// TIA Portal project "Energy_Drink_V15.1" (V15.1) (continued)
REGION Network 3: *****************************MIXER VALVE********************************************/
         A     "Var_System_DB".Sirupe_Valve.Vlv_Open_Cmd;
         =     "Sirupe_Vlv_Man";

         A     "Var_System_DB".Water_Valve.Vlv_Open_Cmd;
         =     "Water_Vlv_Man";

         A     "Var_System_DB".Tk104_MIXER.Open_Vlv_Cmd;
         O     "HMI_VAR".Man_Valves.Mixer_Discharge_Vlv;
         =     "Mixer_Dis_Vlv";

         A     "Var_System_DB".Cleanning_Process.Vlv_Open_Cmd;
         =     "Mixer_Cleanning_Vlv";
END_REGION

REGION Network 4: *****************************CONVEYOR********************************************/
   // CONVEYOR MAIN CONTACTOR
         A     "Var_System_DB".Conveyor_Belt.M_Main;
         =     "KM1_Main";

   // CONVEYOR STAR CONTACTOR
         A     "Var_System_DB".Conveyor_Belt.M_Star;
         =     "KM2_Star";

   // CONVEYOR DELTA CONTACTOR
         A     "Var_System_DB".Conveyor_Belt.M_Led_Delta;
         =     "KM3_Delta";
END_REGION

REGION Network 5: *******************************PROCESS LEDS****************************************/
   // CONVEYOR BELT MOTOR LED ACTIVATION
         A     "Var_System_DB".Conveyor_Belt.M_Led_Main;
         =     "H4";

         A     "Var_System_DB".Conveyor_Belt.M_Led_Delta;
         =     "H5";

         A     "Var_System_DB".Conveyor_Belt.M_Led_Stop;
         =     "H10";

         A     "Var_System_DB".Conveyor_Belt.M_Led_Ovl;
         =     "H8";

   // MIXER MOTOR LED ACTIVATION
         A     "Var_System_DB".Mixer_Motor.Acel_Led;
         =     "H6";

         A     "Var_System_DB".Mixer_Motor.Decel_Led;
         =     "H7";

         A     "Var_System_DB".Mixer_Motor.Led_Ovl;
         =     "H9";
END_REGION
END_FUNCTION

// folder: 02-START-STOP MANGAMENT

FUNCTION "GENERIC_START-STOP" : Void   // FC1, STL
{ S7_Optimized_Access := 'FALSE' }
VERSION : 0.1
BEGIN

REGION Network 1: ******************************* AUTO MODE ********************************************
   // IF START BUTTON PRESSED => DB START
         A     "Start_Button";
         O     "HMI_VAR".Act_System;
         =     "Var_System_DB".System_Generic.Start;

   // IF DB START ACTIVATED => SYSTEM IS ON
         A     "Var_System_DB".System_Generic.Start;
         AN    "Var_System_DB".System_Generic."Auto/Man";
         FP    "Tag_8";
         S     "Var_System_DB".System_Generic.System_Act;
         S     "Var_System_DB".Conveyor_Belt.M_Stop;

   // IF NEGATIVE EDGE OF DB START => RESET
         A     "Var_System_DB".System_Generic.Start;
         FN    "Tag_9";
         R     "Var_System_DB".System_Generic.Stop_Process;
END_REGION

REGION Network 2: ******************************* MANUAL MODE ********************************************
   // SET MANUAL MODE AUTO/MANUAL = 1
         A     "Var_System_DB".System_Generic."Auto/Man";
         A     "Var_System_DB".System_Generic.Start;
         S     "Var_System_DB".System_Generic.Man_Mode;

   // RESET MANUAL MODE
         AN    "Var_System_DB".System_Generic."Auto/Man";
         R     "Var_System_DB".System_Generic.Man_Mode;
END_REGION

REGION Network 3: ******************************* STOP MODE ********************************************
   // WHILE SYSTEM STOP
         A     "Stop_Button";
         A     "HMI_VAR".Stop_System;
         =     "Var_System_DB".System_Generic.Stop;

         AN    "Stop_Button";
         ON    "HMI_VAR".Stop_System;
         S     "Var_System_DB".System_Generic.Stop_Process;
END_REGION
END_FUNCTION

FUNCTION "MOTOR_OVERLOAD_MANAGEMENT" : Void   // FC6, STL
{ S7_Optimized_Access := 'FALSE' }
VERSION : 0.1
BEGIN

REGION Network 1: *************************** SYSTEM FAILURE*****************************************************
         AN    "Var_System_DB".Conveyor_Belt.M_Overload;
         ON    "Var_System_DB".Mixer_Motor.Overload;
         S     "Var_System_DB".System_Generic.System_Failure;

         A     "Var_System_DB".Conveyor_Belt.M_Overload;
         O     "Var_System_DB".Mixer_Motor.Overload;
         A     "Var_System_DB".System_Generic.Start;
         FN    "Tag_25";
         R     "Var_System_DB".System_Generic.System_Failure;
END_REGION
END_FUNCTION

FUNCTION "EMERGENCY_MANGEMENT" : Void   // FC16, STL
{ S7_Optimized_Access := 'FALSE' }
VERSION : 0.1
BEGIN

REGION Network 1: /************************** EMERGENCY STOP MANGEMENT************************************
   // EMERGENCY STOP "NC"
         A     "Emergency_Stop";
         =     "Var_System_DB".System_Generic.Emergency_Stop;

   // IF EMERGENCY STOP IS PRESSED "NA" => RESET ALL
         AN    "Var_System_DB".System_Generic.Emergency_Stop;
         JCN   _800;
         R     "Var_System_DB".System_Generic.System_Act;
         R     "RECIPE_1_DB".Recipe1.Recipe_Act;
         R     "RECIPE_2_DB".Recipe2.Recipe_Act;
         R     "RECIPE_3_DB".Recipe3.Recipe_Act;
         R     "Var_System_DB".System_Generic.Mixer_Station;
         R     "Var_System_DB".Conveyor_Belt.M_Stop;
         R     "Var_System_DB".Mixer_Motor.Motor_Cmd;
         R     "Var_System_DB".Sirupe_Valve.Vlv_Cmd;
         R     "Var_System_DB".Water_Valve.Vlv_Cmd;
         R     "Var_System_DB".System_Generic.Bach_In_Progress;
         R     "Var_System_DB".Conveyor_Belt.State;
         R     "Var_System_DB".Mixer_Motor.State;
         R     "Var_System_DB".Scale_Discharge_Vlv.Vlv_Cmd;
         R     "Var_System_DB".Tk101.Vlv_Cmd;
         R     "Var_System_DB".Tk102.Vlv_Cmd;
         R     "Var_System_DB".Tk103.Vlv_Cmd;
         R     "Var_System_DB".TK101_FILLING_VLV.Vlv_Cmd;
         R     "Var_System_DB".TK102_FILLING_VLV.Vlv_Cmd;
         R     "Var_System_DB".TK103_FILLING_VLV.Vlv_Cmd;

   // SEND THE VALUE "0" TO THE PRODUCTS AND FLOWS SELECTION
         L     0;
         T     "Var_System_DB".Weighing_Process.State;
         T     "M_Product_1";
         T     "M_Product_2";
         T     "M_Product_3";
         T     "M_Water_Flow";
         T     "M_Sirupe_Flow";

   _800: NOP   0;
END_REGION
END_FUNCTION

FUNCTION "START-STOP_MANAGEMENT" : Void   // FC17, FBD
{ S7_Optimized_Access := 'FALSE' }
VERSION : 0.1
BEGIN

REGION Network 1
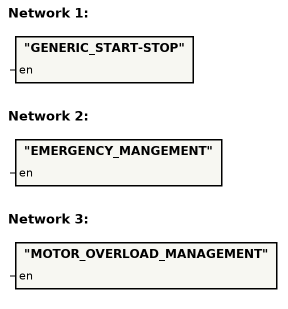
   "GENERIC_START-STOP"();
END_REGION

REGION Network 2
   "EMERGENCY_MANGEMENT"();
END_REGION

REGION Network 3
   "MOTOR_OVERLOAD_MANAGEMENT"();
END_REGION
END_FUNCTION

// folder: 03-TANK MANAGEMENT

FUNCTION "TANKS_MANAGEMENT" : Void   // FC9, FBD
{ S7_Optimized_Access := 'FALSE' }
VERSION : 0.1
BEGIN

REGION Network 1: /************************TANK101 LEVEL *****************************************/
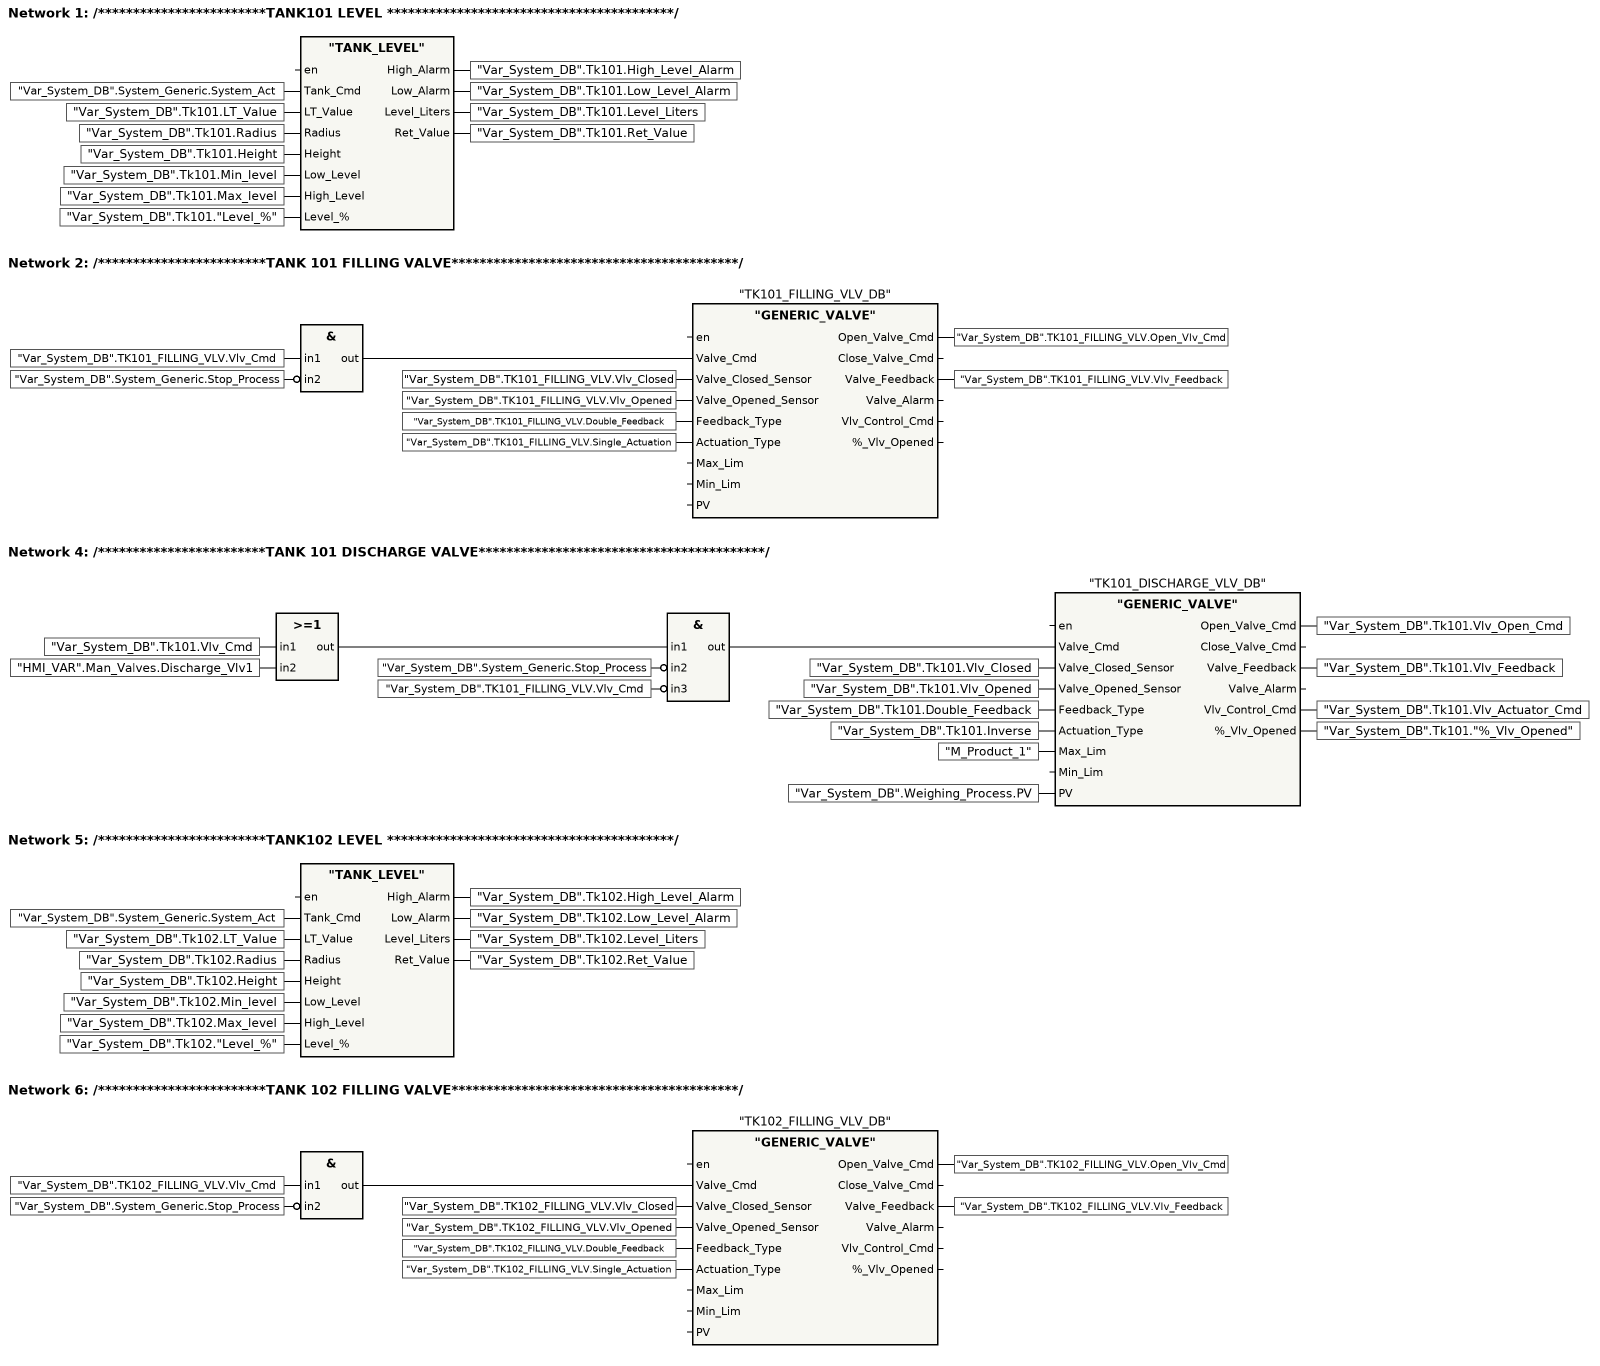
   "TANK_LEVEL"(Tank_Cmd := "Var_System_DB".System_Generic.System_Act,
                LT_Value := "Var_System_DB".Tk101.LT_Value,
                Radius := "Var_System_DB".Tk101.Radius,
                Height := "Var_System_DB".Tk101.Height,
                Low_Level := "Var_System_DB".Tk101.Min_level,
                High_Level := "Var_System_DB".Tk101.Max_level,
                "Level_%" := "Var_System_DB".Tk101."Level_%",
                High_Alarm => "Var_System_DB".Tk101.High_Level_Alarm,
                Low_Alarm => "Var_System_DB".Tk101.Low_Level_Alarm,
                Level_Liters => "Var_System_DB".Tk101.Level_Liters,
                Ret_Value => "Var_System_DB".Tk101.Ret_Value);
END_REGION

REGION Network 2: /************************TANK 101 FILLING VALVE*****************************************/
   "TK101_FILLING_VLV_DB"(Valve_Cmd := "Var_System_DB".TK101_FILLING_VLV.Vlv_Cmd AND NOT "Var_System_DB".System_Generic.Stop_Process,   // "GENERIC_VALVE"
                          Valve_Closed_Sensor := "Var_System_DB".TK101_FILLING_VLV.Vlv_Closed,
                          Valve_Opened_Sensor := "Var_System_DB".TK101_FILLING_VLV.Vlv_Opened,
                          Feedback_Type := "Var_System_DB".TK101_FILLING_VLV.Double_Feedback,
                          Actuation_Type := "Var_System_DB".TK101_FILLING_VLV.Single_Actuation,
                          Open_Valve_Cmd => "Var_System_DB".TK101_FILLING_VLV.Open_Vlv_Cmd,
                          Valve_Feedback => "Var_System_DB".TK101_FILLING_VLV.Vlv_Feedback);
END_REGION

REGION Network 3 (STL): ************************CONDITIONS TO FILL TANK 101*****************************************/
   // IF SYSTEM IS ACTIVE => CHECK CONDITIONS
         A     "Var_System_DB".System_Generic.System_Act;
   // IF LEVEL IS < 20% => SET FILLING TANK
         A(;
         L     "Var_System_DB".Tk101."Level_%";
         L     20;
         <=I;
         );
         S     "Var_System_DB".TK101_FILLING_VLV.Vlv_Cmd;  // SET VLV_CMD

   // IF LEVEL IS >= 90% => RESET FILLING TANK
         A(;
         L     "Var_System_DB".Tk101."Level_%";
         L     90;
         >=I;
         );
         R     "Var_System_DB".TK101_FILLING_VLV.Vlv_Cmd;  // RESET VLV_CMD
END_REGION

REGION Network 4: /************************TANK 101 DISCHARGE VALVE*****************************************/
   "TK101_DISCHARGE_VLV_DB"(Valve_Cmd := ("Var_System_DB".Tk101.Vlv_Cmd OR "HMI_VAR".Man_Valves.Discharge_Vlv1) AND NOT "Var_System_DB".System_Generic.Stop_Process AND NOT "Var_System_DB".TK101_FILLING_VLV.Vlv_Cmd,   // "GENERIC_VALVE"
                           Valve_Closed_Sensor := "Var_System_DB".Tk101.Vlv_Closed,
                           Valve_Opened_Sensor := "Var_System_DB".Tk101.Vlv_Opened,
                           Feedback_Type := "Var_System_DB".Tk101.Double_Feedback,
                           Actuation_Type := "Var_System_DB".Tk101.Inverse,
                           Max_Lim := "M_Product_1",
                           PV := "Var_System_DB".Weighing_Process.PV,
                           Open_Valve_Cmd => "Var_System_DB".Tk101.Vlv_Open_Cmd,
                           Valve_Feedback => "Var_System_DB".Tk101.Vlv_Feedback,
                           Vlv_Control_Cmd => "Var_System_DB".Tk101.Vlv_Actuator_Cmd,
                           "%_Vlv_Opened" => "Var_System_DB".Tk101."%_Vlv_Opened");
END_REGION

REGION Network 5: /************************TANK102 LEVEL *****************************************/
   "TANK_LEVEL"(Tank_Cmd := "Var_System_DB".System_Generic.System_Act,
                LT_Value := "Var_System_DB".Tk102.LT_Value,
                Radius := "Var_System_DB".Tk102.Radius,
                Height := "Var_System_DB".Tk102.Height,
                Low_Level := "Var_System_DB".Tk102.Min_level,
                High_Level := "Var_System_DB".Tk102.Max_level,
                "Level_%" := "Var_System_DB".Tk102."Level_%",
                High_Alarm => "Var_System_DB".Tk102.High_Level_Alarm,
                Low_Alarm => "Var_System_DB".Tk102.Low_Level_Alarm,
                Level_Liters => "Var_System_DB".Tk102.Level_Liters,
                Ret_Value => "Var_System_DB".Tk102.Ret_Value);
END_REGION

REGION Network 6: /************************TANK 102 FILLING VALVE*****************************************/
   "TK102_FILLING_VLV_DB"(Valve_Cmd := "Var_System_DB".TK102_FILLING_VLV.Vlv_Cmd AND NOT "Var_System_DB".System_Generic.Stop_Process,   // "GENERIC_VALVE"
                          Valve_Closed_Sensor := "Var_System_DB".TK102_FILLING_VLV.Vlv_Closed,
                          Valve_Opened_Sensor := "Var_System_DB".TK102_FILLING_VLV.Vlv_Opened,
                          Feedback_Type := "Var_System_DB".TK102_FILLING_VLV.Double_Feedback,
                          Actuation_Type := "Var_System_DB".TK102_FILLING_VLV.Single_Actuation,
                          Open_Valve_Cmd => "Var_System_DB".TK102_FILLING_VLV.Open_Vlv_Cmd,
                          Valve_Feedback => "Var_System_DB".TK102_FILLING_VLV.Vlv_Feedback);
END_REGION

REGION Network 7 (STL): ************************CONDITIONS TO FILL TANK 102*****************************************/
   // IF SYSTEM IS ACTIVE => CHECK CONDITIONS
         A     "Var_System_DB".System_Generic.System_Act;
   // IF LEVEL IS < 20% => SET FILLING TANK
         A(;
         L     "Var_System_DB".Tk102."Level_%";
         L     20;
         <=I;
         );
         S     "Var_System_DB".TK102_FILLING_VLV.Vlv_Cmd;  // SET VLV_CMD

   // IF LEVEL IS >= 90% => RESET FILLING TANK
         A(;
         L     "Var_System_DB".Tk102."Level_%";
         L     90;
         >=I;
         );
         R     "Var_System_DB".TK102_FILLING_VLV.Vlv_Cmd;  // RESET VLV_CMD
END_REGION

REGION Network 8 (STL): /************************DISCHARGE VLV 2 MAX LIMIT*****************************************/
   // SUM OF THE PRODUCT 1 AND 2 TO USE IT AS A MAX LIMIT FOR DISCHARGE VLV 2
         L     "M_Product_1";
         L     "M_Product_2";
         +R;
         T     "Temp_Lim_Kg";  // DISCHARGE VLV 2 MAX LIMIT
END_REGION

REGION Network 9: /************************TANK 102 AND DISCHARGE VALVE*****************************************/
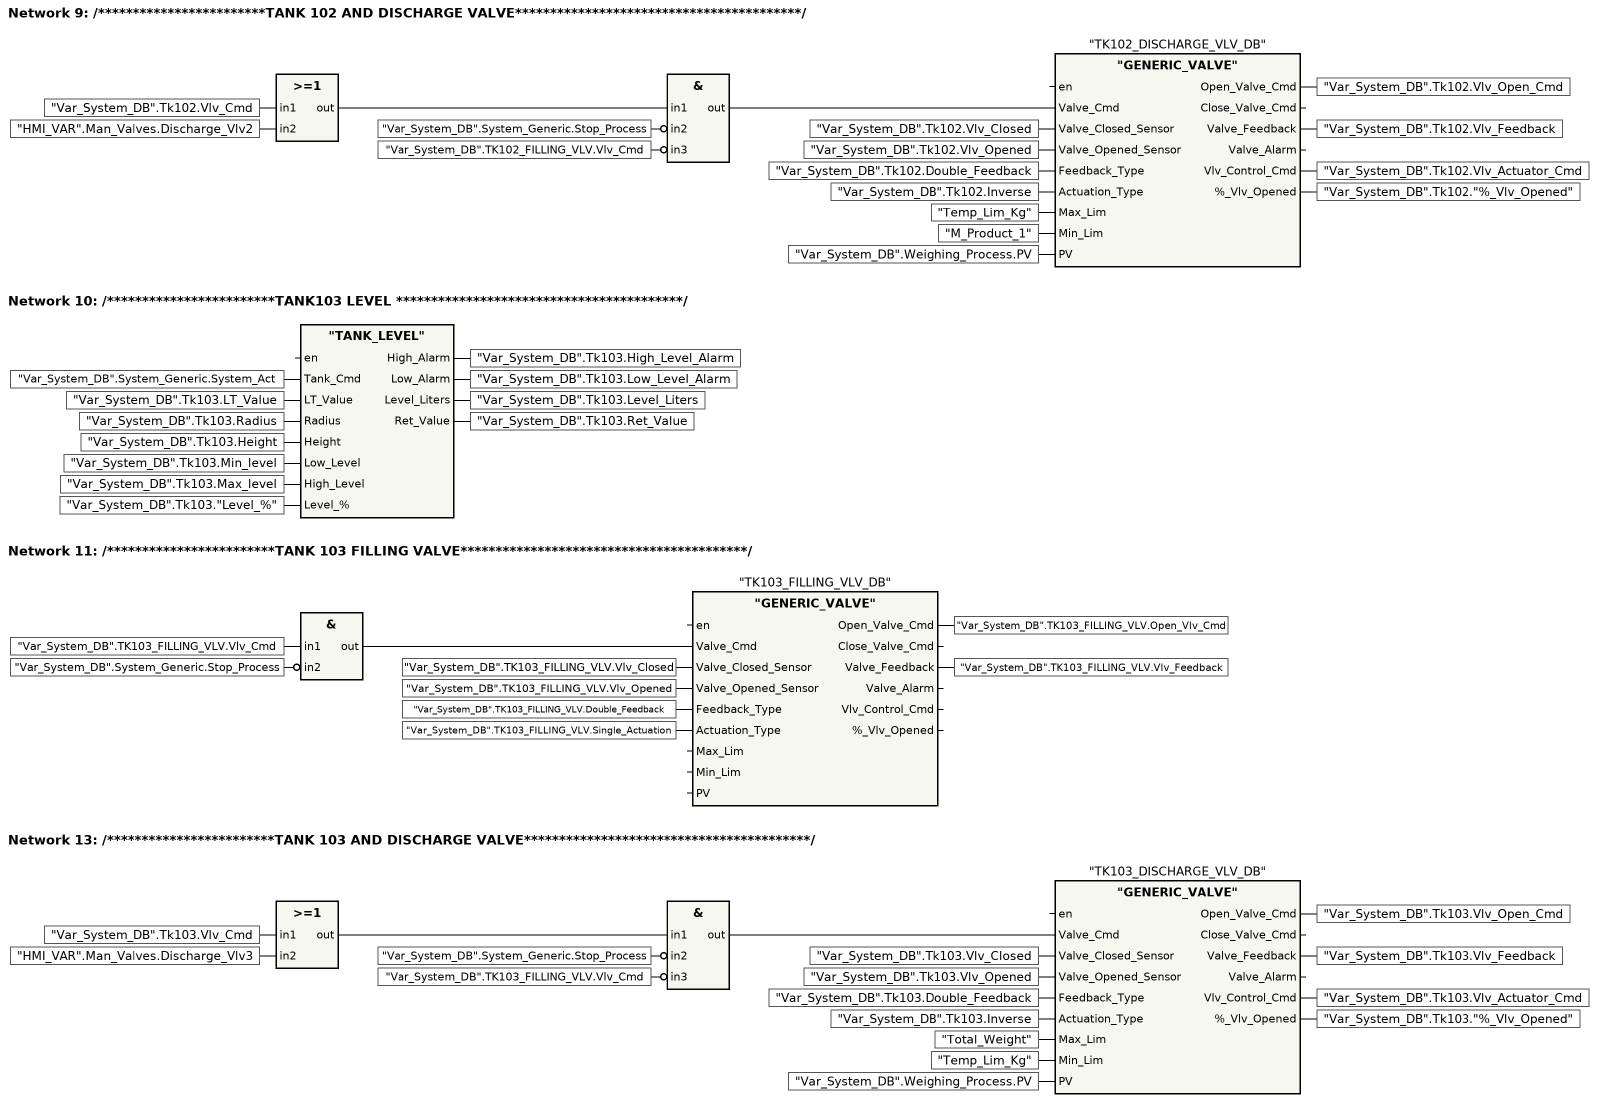
   "TK102_DISCHARGE_VLV_DB"(Valve_Cmd := ("Var_System_DB".Tk102.Vlv_Cmd OR "HMI_VAR".Man_Valves.Discharge_Vlv2) AND NOT "Var_System_DB".System_Generic.Stop_Process AND NOT "Var_System_DB".TK102_FILLING_VLV.Vlv_Cmd,   // "GENERIC_VALVE"
                           Valve_Closed_Sensor := "Var_System_DB".Tk102.Vlv_Closed,
                           Valve_Opened_Sensor := "Var_System_DB".Tk102.Vlv_Opened,
                           Feedback_Type := "Var_System_DB".Tk102.Double_Feedback,
                           Actuation_Type := "Var_System_DB".Tk102.Inverse,
                           Max_Lim := "Temp_Lim_Kg",
                           Min_Lim := "M_Product_1",
                           PV := "Var_System_DB".Weighing_Process.PV,
                           Open_Valve_Cmd => "Var_System_DB".Tk102.Vlv_Open_Cmd,
                           Valve_Feedback => "Var_System_DB".Tk102.Vlv_Feedback,
                           Vlv_Control_Cmd => "Var_System_DB".Tk102.Vlv_Actuator_Cmd,
                           "%_Vlv_Opened" => "Var_System_DB".Tk102."%_Vlv_Opened");
END_REGION

REGION Network 10: /************************TANK103 LEVEL *****************************************/
   "TANK_LEVEL"(Tank_Cmd := "Var_System_DB".System_Generic.System_Act,
                LT_Value := "Var_System_DB".Tk103.LT_Value,
                Radius := "Var_System_DB".Tk103.Radius,
                Height := "Var_System_DB".Tk103.Height,
                Low_Level := "Var_System_DB".Tk103.Min_level,
                High_Level := "Var_System_DB".Tk103.Max_level,
                "Level_%" := "Var_System_DB".Tk103."Level_%",
                High_Alarm => "Var_System_DB".Tk103.High_Level_Alarm,
                Low_Alarm => "Var_System_DB".Tk103.Low_Level_Alarm,
                Level_Liters => "Var_System_DB".Tk103.Level_Liters,
                Ret_Value => "Var_System_DB".Tk103.Ret_Value);
END_REGION

REGION Network 11: /************************TANK 103 FILLING VALVE*****************************************/
   "TK103_FILLING_VLV_DB"(Valve_Cmd := "Var_System_DB".TK103_FILLING_VLV.Vlv_Cmd AND NOT "Var_System_DB".System_Generic.Stop_Process,   // "GENERIC_VALVE"
                          Valve_Closed_Sensor := "Var_System_DB".TK103_FILLING_VLV.Vlv_Closed,
                          Valve_Opened_Sensor := "Var_System_DB".TK103_FILLING_VLV.Vlv_Opened,
                          Feedback_Type := "Var_System_DB".TK103_FILLING_VLV.Double_Feedback,
                          Actuation_Type := "Var_System_DB".TK103_FILLING_VLV.Single_Actuation,
                          Open_Valve_Cmd => "Var_System_DB".TK103_FILLING_VLV.Open_Vlv_Cmd,
                          Valve_Feedback => "Var_System_DB".TK103_FILLING_VLV.Vlv_Feedback);
END_REGION

REGION Network 12 (STL): ************************CONDITIONS TO FILL TANK 103*****************************************/
   // IF SYSTEM IS ACTIVE => CHECK CONDITIONS
         A     "Var_System_DB".System_Generic.System_Act;
   // IF LEVEL IS < 20% => SET FILLING TANK
         A(;
         L     "Var_System_DB".Tk103."Level_%";
         L     20;
         <=I;
         );
         S     "Var_System_DB".TK103_FILLING_VLV.Vlv_Cmd;  // SET VLV_CMD

   // IF LEVEL IS >= 90% => RESET FILLING TANK
         A(;
         L     "Var_System_DB".Tk103."Level_%";
         L     90;
         >=I;
         );
         R     "Var_System_DB".TK103_FILLING_VLV.Vlv_Cmd;  // RESET VLV_CMD
END_REGION

REGION Network 13: /************************TANK 103 AND DISCHARGE VALVE*****************************************/
   "TK103_DISCHARGE_VLV_DB"(Valve_Cmd := ("Var_System_DB".Tk103.Vlv_Cmd OR "HMI_VAR".Man_Valves.Discharge_Vlv3) AND NOT "Var_System_DB".System_Generic.Stop_Process AND NOT "Var_System_DB".TK103_FILLING_VLV.Vlv_Cmd,   // "GENERIC_VALVE"
                           Valve_Closed_Sensor := "Var_System_DB".Tk103.Vlv_Closed,
                           Valve_Opened_Sensor := "Var_System_DB".Tk103.Vlv_Opened,
                           Feedback_Type := "Var_System_DB".Tk103.Double_Feedback,
                           Actuation_Type := "Var_System_DB".Tk103.Inverse,
                           Max_Lim := "Total_Weight",
                           Min_Lim := "Temp_Lim_Kg",
                           PV := "Var_System_DB".Weighing_Process.PV,
                           Open_Valve_Cmd => "Var_System_DB".Tk103.Vlv_Open_Cmd,
                           Valve_Feedback => "Var_System_DB".Tk103.Vlv_Feedback,
                           Vlv_Control_Cmd => "Var_System_DB".Tk103.Vlv_Actuator_Cmd,
                           "%_Vlv_Opened" => "Var_System_DB".Tk103."%_Vlv_Opened");
END_REGION
END_FUNCTION

// folder: 04-OPERATOR MANAGEMENT

FUNCTION "PROD_WEIGHING_MANAGEMENT" : Void   // FC4, STL
{ S7_Optimized_Access := 'FALSE' }
VERSION : 0.1
   VAR_INPUT
      Product_1 : Real;
      Product_2 : Real;
      Product_3 : Real;
      Water_Flow : Real;
      Sirupe_Flow : Real;
      Num_Bach : Int;   // Number of batches to produce
   END_VAR
   VAR_TEMP
      Weight_Kg : Real;
   END_VAR
BEGIN

REGION Network 1: /************************MAPPING OF INPUT PARAMETERS *****************************************/
   // DUE TO THE AUF COMMAND FROM FC "RECIPE SELECTION"
   // MAPPING INPUTS FROM DB PARAMETERS => MEMORY VAR
         L     #Product_1;
         T     "M_Product_1";
         L     #Product_2;
         T     "M_Product_2";
         L     #Product_3;
         T     "M_Product_3";
         L     #Water_Flow;
         T     "M_Water_Flow";
         L     #Sirupe_Flow;
         T     "M_Sirupe_Flow";
         L     #Num_Bach;
         T     "Num_Bach";

   // CALCULATE TOTAL WEIGHT IN KG
         L     "M_Product_1";
         L     "M_Product_2";
         +R;
         L     "M_Product_3";
         +R;
         T     "Total_Weight";

   // IF RESET BUTTON PRESSED LOAD "0" TO WEIGHT_KG
         A     "Reset_Button";
         JCN   _305;
         L     0;
         T     #Weight_Kg;
   _305: NOP   0;
END_REGION

REGION Network 2: /************************ SCALING SENSOR ACTIVATION *****************************************/
   // SCALE SENSOR
         CALL  SCALE
         ( IN      := "Weighing":P,
           HI_LIM  := "Var_System_DB".Weighing_Process.Max_Kg,
           LO_LIM  := "Var_System_DB".Weighing_Process.Min_Kg,
           BIPOLAR := FALSE,
           RET_VAL := "Recipe_Num",
           OUT     := "Var_System_DB".Weighing_Process.PV
         );


   // MOVE PROCESS VARIABLE PV => WEIGHT_KG
         L     "Var_System_DB".Weighing_Process.PV;
         T     #Weight_Kg;
END_REGION

REGION Network 3: /************************CONDITIONS TO OPEN TANK VALVES *****************************************/
   // IF NOT BACH IN PROGRESS
         A     "HMI_VAR".Start_Process;
         O     "Var_System_DB".System_Generic.Man_Start_Process;
         AN    "Var_System_DB".System_Generic.Bach_In_Progress;
         JCN   _300;
         L     "Var_System_DB".Weighing_Process.State;  // VAR TO MANAGE THE JUMPS TO THE DIFFERENT WEIGHING STATES

   // CASE STATEMENT TO PERFORM AND ACTION BASED ON STAGE OF THE PROCESS
         JL    _301;

         JU    PROD1;  // IF "0" GO TO PROD1
         JU    PROD2;  // IF "1" GO TO PROD2
         JU    PROD3;  // IF "2" GO TO PROD3

   _301: JU    OUT;

   // PRODUCT 1 CONDITIONS TO SEND COMMAND TO OPEN TANK 1 DISCHARGE  VALVE
   PROD1:A(;
         L     #Weight_Kg;
         L     "M_Product_1";
         <R;
         );
         =     "Var_System_DB".Tk101.Vlv_Cmd;  // SEND COMMAND TO OPEN TANK 101 DISCHARGE VALVE

   // IF WEIGTH >= PROCESS_STATE  = 1, GO TO NEXT TANK
         A(;
         L     #Weight_Kg;
         L     "M_Product_1";
         >=R;
         );
         JCN   _302;
         L     1;
         T     "Var_System_DB".Weighing_Process.State;  // MODIFY VALUE TO GO TO THE NEXT WEIGHING STATE
   _302: NOP   0;
         JU    END;

   // PRODUCT 2 CONDITIONS TO SEND COMMAND TO OPEN TANK 2 DISCHARGE  VALVE
   PROD2:A(;
         L     "M_Product_1";
         L     "M_Product_2";
         +R;
         L     #Weight_Kg;
         >R;
         );
         =     "Var_System_DB".Tk102.Vlv_Cmd;  // SEND COMMAND TO OPEN TANK 102 DISCHARGE VALVE

   // IF WEIGTH >= PROCESS_STATE  = 1, GO TO NEXT TANK
         A(;
         L     "M_Product_1";
         L     "M_Product_2";
         +R;
         L     #Weight_Kg;
         <=R;
         );
         JCN   _303;
         L     2;
         T     "Var_System_DB".Weighing_Process.State;  // MODIFY VALUE TO GO TO FINAL WEIGHING STATE
   _303: NOP   0;

         JU    END;


   // PRODUCT 3 CONDITIONS TO SEND COMMAND TO OPEN TANK 3 DISCHARGE  VALVE
   PROD3:A(;
         L     "M_Product_1";
         L     "M_Product_2";
         +R;
         L     "M_Product_3";
         +R;
         L     #Weight_Kg;
         >R;
         );
         =     "Var_System_DB".Tk103.Vlv_Cmd;  // SEND COMMAND TO OPEN TANK 103 DISCHARGE VALVE

   // IF WEIGTH >= SCALE_PV => PROCESS_STATE  = 0 => BACH IN PROCESS ACTIVE
         A(;
         L     "M_Product_1";
         L     "M_Product_2";
         +R;
         L     "M_Product_3";
         +R;
         L     #Weight_Kg;
         <=R;
         );
         JCN   _304;
         S     "Var_System_DB".System_Generic.Bach_In_Progress;
         L     0;
         T     "Var_System_DB".Weighing_Process.State;  // // RESET VALUE TO ITS INITIAL STAT
   _304: NOP   0;

         JU    END;

   // IF VALUE OUT OF RANGE => SET PROCESS_STATE = 0 (INITIAL VALUE)
   OUT:  L     0;
         T     "Var_System_DB".Weighing_Process.State;

         JU    END;

   // IF JUMPED TO END GET OUT OF THE LOOP
   END:  BEU;

   _300: NOP   0;
END_REGION

REGION Network 4: /************************SCALE DISCHARGE VALVE *****************************************/
   // WHILE THE SCALE SENSOR IS GREATER THAN "0" KG
         A     "Var_System_DB".System_Generic.Bach_In_Progress;
         A(;
         L     #Weight_Kg;
         L     0;
         >R;
         );
         =     "Var_System_DB".Scale_Discharge_Vlv.Vlv_Cmd;  // SEND COMMAND TO OPEN SCALE DISCAHRGE VALVE


   // WHILE THE CONDITION ARE MET => SEND COMMAND TO OPEN THE VALE
         A     "Var_System_DB".Scale_Discharge_Vlv.Vlv_Cmd;
         A     "Var_System_DB".System_Generic.Stop;
         =     "Var_System_DB".Scale_Discharge_Vlv.Open_Vlv_Cmd;


   // FB GENERIC VALVE CALL
         CALL  "GENERIC_VALVE", "SCALE_DISCHARGE_VLV_DB"
         ( Valve_Cmd           := "Var_System_DB".Scale_Discharge_Vlv.Open_Vlv_Cmd,
           Valve_Closed_Sensor := "Var_System_DB".Scale_Discharge_Vlv.Vlv_Closed,
           Valve_Opened_Sensor := "Var_System_DB".Scale_Discharge_Vlv.Vlv_Opened,
           Feedback_Type       := "Var_System_DB".Scale_Discharge_Vlv.Double_Feedback,
           Actuation_Type      := "Var_System_DB".Scale_Discharge_Vlv.Single_Actuation,
           Max_Lim             := ,
           Min_Lim             := ,
           PV                  := ,
           Open_Valve_Cmd      := "Var_System_DB".Scale_Discharge_Vlv.Open_Vlv,
           Close_Valve_Cmd     := ,
           Valve_Feedback      := "Var_System_DB".Scale_Discharge_Vlv.Vlv_Feedback,
           Valve_Alarm         := ,
           Vlv_Control_Cmd     := ,
           "%_Vlv_Opened"      :=
         );
END_REGION
END_FUNCTION

FUNCTION "RECIPE_MANAGEMENT" : Void   // FC11, STL
{ S7_Optimized_Access := 'FALSE' }
VERSION : 0.1
BEGIN

REGION Network 1: *********************CHECK OPERATORS SELECTIONS*************************************
   // IF THE SYSTEM IS ACTIVE AND NOT MIXER_STATION AND RECIPE_ACT
   // CHECK THE NUMBER OF "RECIPE" TO OPEN THE CORRESPONDING DB
         A     "Var_System_DB".System_Generic.System_Act;
         A(;
         A     "RECIPE_1_DB".Recipe1.Recipe_Act;
         O     "RECIPE_2_DB".Recipe2.Recipe_Act;
         O     "RECIPE_3_DB".Recipe3.Recipe_Act;
         O     "TEST_RECIPE_DB".Test.Recipe_Act;
         );
         A(;
         L     "Recipe_Num";
         L     10;
         >=I;
         );
         A(;
         L     "Recipe_Num";
         L     13;
         <=I;
         );
         JCN   _200;
   // IF THE VALUE OF RECIPE_NUM IS BETWEEN 10-13 => OPEN DB[RECIPE_NUMBER]
   // CALL "FC PRODUCTS WEIGNING MANAGEMENT" WITH THE CORRESPONDING PARAMETERS FROM DB

         OPN   DB [ "Recipe_Num"];

         CALL  "PROD_WEIGHING_MANAGEMENT"
         ( Product_1   := %DataD4,
           Product_2   := %DataD8,
           Product_3   := %DataD12,
           Water_Flow  := %DataD16,
           Sirupe_Flow := %DataD20,
           Num_Bach    := %DataW2
         );

   _200: NOP   0;
END_REGION
END_FUNCTION

FUNCTION "OP_RECIPE_SELCT" : Void   // FC12, SCL
{ S7_Optimized_Access := 'FALSE' }
VERSION : 0.1
BEGIN
   (*
   *File: FC Operator Recipe Selection
   * Author: Jaime Calvente Mieres
   * Date: 19-05-2022
   * Description: This FC will be used to control a valve. Depending on 
     the users input, the valve could act as Single actuation,
     Double actuation or Proportional mode.
   *)

   // RECIPE MANAGEMENT CALL
   "RECIPE_MANAGEMENT"();

   (************************ SET RECIPE SELECTION MANAGEMENT **********************************)
   REGION SET RECIPE SELECTION

       // IF SYSTEM IS ACTIVE WAIT FOR THE OPERATOR TO CHOOSE THE RECIPE BY HMI OR CONTOL PANEL "MANUAL"
       IF "Var_System_DB".System_Generic.System_Act THEN

           // IF NOT RECIPE ACTIVE
           "Var_System_DB".System_Generic.No_Process := NOT "RECIPE_1_DB".Recipe1.Recipe_Act AND
           NOT "RECIPE_2_DB".Recipe2.Recipe_Act AND
           NOT "RECIPE_3_DB".Recipe3.Recipe_Act AND
           NOT "TEST_RECIPE_DB".Test.Recipe_Act;

           (*This Nested If statements will be executed only if the System is
           Active and there is NO bacth in process, checking the variable 
           "No_Process" and the Operator selection  (switches or HMI).*)

           REGION RECIPE SELECTION

               // IF NOT ACTIVE PROCESS
               IF "Var_System_DB".System_Generic.No_Process THEN

                   // IF RECIPE NUMBER 1 => SET "RECIPE_1_DB"   
                   IF "Recipe_1" OR "HMI_VAR".Recipe_Selection[1] THEN
                       "RECIPE_1_DB".Recipe1.Recipe_Act := TRUE;
                   ELSIF "Recipe_2" OR "Recipe_3" THEN
                       "RECIPE_1_DB".Recipe1.Recipe_Act := FALSE;
                   END_IF;


                   // IF RECIPE NUMBER 2 => SET "RECIPE_2_DB"   
                   IF "Recipe_2" OR "HMI_VAR".Recipe_Selection[2] THEN
                       "RECIPE_2_DB".Recipe2.Recipe_Act := TRUE;
                   ELSIF "Recipe_1" OR "Recipe_3" THEN
                       "RECIPE_2_DB".Recipe2.Recipe_Act := FALSE;
                   END_IF;

                   // IF RECIPE NUMBER 3 => SET "RECIPE_3_DB"     
                   IF "Recipe_3" OR "HMI_VAR".Recipe_Selection[3] THEN
                       "RECIPE_3_DB".Recipe3.Recipe_Act := TRUE;
                   ELSIF "Recipe_1" OR "Recipe_2" THEN
                       "RECIPE_3_DB".Recipe3.Recipe_Act := FALSE;
                   END_IF;

                   // TEST RECIPE
                   IF "HMI_VAR".Recipe_Selection[4] THEN
                       "TEST_RECIPE_DB".Test.Recipe_Act := TRUE;
                   ELSIF "Recipe_1" OR "Recipe_2" OR "Recipe_3" THEN
                       "TEST_RECIPE_DB".Test.Recipe_Act := FALSE;
                   END_IF;
               END_IF;

           END_REGION

           (*This Nested IF statement will set the Variable "Recipe_Num" TO 
            a value according TO the specific DB number needed in order TO 
            access the parameters OF the chosen Recipe.*)

           REGION RECIPE NUMBER FOR DB SELECTION

               // IF "RECIPE_1_DB"  => "Recipe_Num" = 10
               IF "RECIPE_1_DB".Recipe1.Recipe_Act THEN
                   "Recipe_Num" := 10;
               END_IF;

               // IF "RECIPE_2_DB"  => RECIPE_NUM = 11
               IF "RECIPE_2_DB".Recipe2.Recipe_Act THEN
                   "Recipe_Num" := 11;
               END_IF;

               // IF "RECIPE_3_DB"  => "Recipe_Num" = 12
               IF "RECIPE_3_DB".Recipe3.Recipe_Act THEN
                   "Recipe_Num" := 12;
               END_IF;

               // IF "RECIPE_TEST"  => "Recipe_Num" = 13
               IF "TEST_RECIPE_DB".Test.Recipe_Act THEN
                   "Recipe_Num" := 13;
               END_IF;

           END_REGION

       // IF SYSTEM IS NOT ACTIVE => NOT RECIPE WILL BE SELECTED RETURNING THE VALUE OF "0"    
       ELSE
           "RECIPE_1_DB".Recipe1.Recipe_Act := FALSE;
           "RECIPE_2_DB".Recipe2.Recipe_Act := FALSE;
           "RECIPE_3_DB".Recipe3.Recipe_Act := FALSE;
           "TEST_RECIPE_DB".Test.Recipe_Act := FALSE;
           "Recipe_Num" := 0;
           "Var_System_DB".System_Generic.Man_Start_Process := FALSE;
           "HMI_VAR".Start_Process := FALSE;

       END_IF;

   END_REGION

   (************************ RESET RECIPE SELECTION MANAGEMENT **********************************)
   REGION  RESET RECIPE SELECTION